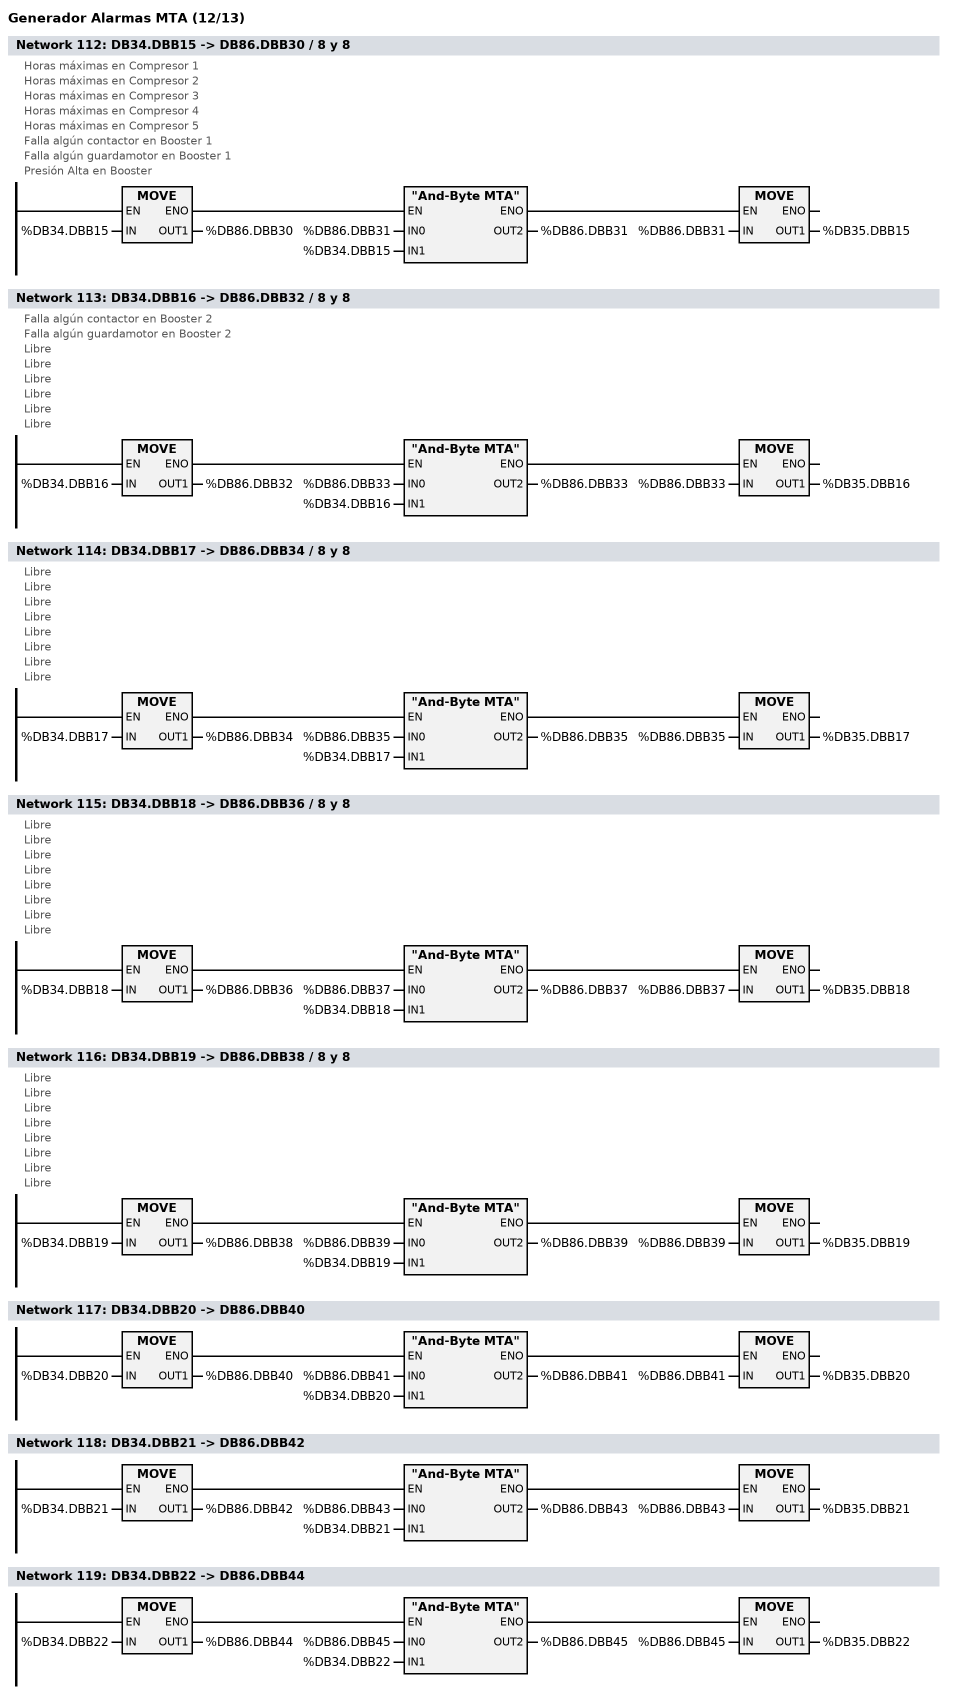
   RUNG wire#powerrail
      { S7_GenerateENO := "TRUE" } Move(in := %DB34.DBB15, out1 => %DB86.DBB30)
      "And-Byte MTA"(IN0 := %DB86.DBB31, IN1 := %DB34.DBB15, OUT2 => %DB86.DBB31)
      { S7_GenerateENO := "TRUE" } Move(in := %DB86.DBB31, out1 => %DB35.DBB15)
   END_RUNG
   // the same network as SCL:
   // ENO of a box is taken as its EN; it also drops when the box reports an error
   %DB86.DBB30 := %DB34.DBB15;
   "And-Byte MTA"(IN0 := %DB86.DBB31, IN1 := %DB34.DBB15, OUT2 => %DB86.DBB31, ENO => #_w1);
   IF #_w1 THEN %DB35.DBB15 := %DB86.DBB31; END_IF;
END_REGION

REGION Network 113: DB34.DBB16 -> DB86.DBB32 / 8 y 8
   // Falla algún contactor en Booster 2
   // Falla algún guardamotor en Booster 2
   // Libre
   // Libre
   // Libre
   // Libre
   // Libre
   // Libre
   RUNG wire#powerrail
      { S7_GenerateENO := "TRUE" } Move(in := %DB34.DBB16, out1 => %DB86.DBB32)
      "And-Byte MTA"(IN0 := %DB86.DBB33, IN1 := %DB34.DBB16, OUT2 => %DB86.DBB33)
      { S7_GenerateENO := "TRUE" } Move(in := %DB86.DBB33, out1 => %DB35.DBB16)
   END_RUNG
   // the same network as SCL:
   // ENO of a box is taken as its EN; it also drops when the box reports an error
   %DB86.DBB32 := %DB34.DBB16;
   "And-Byte MTA"(IN0 := %DB86.DBB33, IN1 := %DB34.DBB16, OUT2 => %DB86.DBB33, ENO => #_w1);
   IF #_w1 THEN %DB35.DBB16 := %DB86.DBB33; END_IF;
END_REGION

REGION Network 114: DB34.DBB17 -> DB86.DBB34 / 8 y 8
   // Libre
   // Libre
   // Libre
   // Libre
   // Libre
   // Libre
   // Libre
   // Libre
   RUNG wire#powerrail
      { S7_GenerateENO := "TRUE" } Move(in := %DB34.DBB17, out1 => %DB86.DBB34)
      "And-Byte MTA"(IN0 := %DB86.DBB35, IN1 := %DB34.DBB17, OUT2 => %DB86.DBB35)
      { S7_GenerateENO := "TRUE" } Move(in := %DB86.DBB35, out1 => %DB35.DBB17)
   END_RUNG
   // the same network as SCL:
   // ENO of a box is taken as its EN; it also drops when the box reports an error
   %DB86.DBB34 := %DB34.DBB17;
   "And-Byte MTA"(IN0 := %DB86.DBB35, IN1 := %DB34.DBB17, OUT2 => %DB86.DBB35, ENO => #_w1);
   IF #_w1 THEN %DB35.DBB17 := %DB86.DBB35; END_IF;
END_REGION

REGION Network 115: DB34.DBB18 -> DB86.DBB36 / 8 y 8
   // Libre
   // Libre
   // Libre
   // Libre
   // Libre
   // Libre
   // Libre
   // Libre
   RUNG wire#powerrail
      { S7_GenerateENO := "TRUE" } Move(in := %DB34.DBB18, out1 => %DB86.DBB36)
      "And-Byte MTA"(IN0 := %DB86.DBB37, IN1 := %DB34.DBB18, OUT2 => %DB86.DBB37)
      { S7_GenerateENO := "TRUE" } Move(in := %DB86.DBB37, out1 => %DB35.DBB18)
   END_RUNG
   // the same network as SCL:
   // ENO of a box is taken as its EN; it also drops when the box reports an error
   %DB86.DBB36 := %DB34.DBB18;
   "And-Byte MTA"(IN0 := %DB86.DBB37, IN1 := %DB34.DBB18, OUT2 => %DB86.DBB37, ENO => #_w1);
   IF #_w1 THEN %DB35.DBB18 := %DB86.DBB37; END_IF;
END_REGION

REGION Network 116: DB34.DBB19 -> DB86.DBB38 / 8 y 8
   // Libre
   // Libre
   // Libre
   // Libre
   // Libre
   // Libre
   // Libre
   // Libre
   RUNG wire#powerrail
      { S7_GenerateENO := "TRUE" } Move(in := %DB34.DBB19, out1 => %DB86.DBB38)
      "And-Byte MTA"(IN0 := %DB86.DBB39, IN1 := %DB34.DBB19, OUT2 => %DB86.DBB39)
      { S7_GenerateENO := "TRUE" } Move(in := %DB86.DBB39, out1 => %DB35.DBB19)
   END_RUNG
   // the same network as SCL:
   // ENO of a box is taken as its EN; it also drops when the box reports an error
   %DB86.DBB38 := %DB34.DBB19;
   "And-Byte MTA"(IN0 := %DB86.DBB39, IN1 := %DB34.DBB19, OUT2 => %DB86.DBB39, ENO => #_w1);
   IF #_w1 THEN %DB35.DBB19 := %DB86.DBB39; END_IF;
END_REGION

REGION Network 117: DB34.DBB20 -> DB86.DBB40
   RUNG wire#powerrail
      { S7_GenerateENO := "TRUE" } Move(in := %DB34.DBB20, out1 => %DB86.DBB40)
      "And-Byte MTA"(IN0 := %DB86.DBB41, IN1 := %DB34.DBB20, OUT2 => %DB86.DBB41)
      { S7_GenerateENO := "TRUE" } Move(in := %DB86.DBB41, out1 => %DB35.DBB20)
   END_RUNG
   // the same network as SCL:
   // ENO of a box is taken as its EN; it also drops when the box reports an error
   %DB86.DBB40 := %DB34.DBB20;
   "And-Byte MTA"(IN0 := %DB86.DBB41, IN1 := %DB34.DBB20, OUT2 => %DB86.DBB41, ENO => #_w1);
   IF #_w1 THEN %DB35.DBB20 := %DB86.DBB41; END_IF;
END_REGION

REGION Network 118: DB34.DBB21 -> DB86.DBB42
   RUNG wire#powerrail
      { S7_GenerateENO := "TRUE" } Move(in := %DB34.DBB21, out1 => %DB86.DBB42)
      "And-Byte MTA"(IN0 := %DB86.DBB43, IN1 := %DB34.DBB21, OUT2 => %DB86.DBB43)
      { S7_GenerateENO := "TRUE" } Move(in := %DB86.DBB43, out1 => %DB35.DBB21)
   END_RUNG
   // the same network as SCL:
   // ENO of a box is taken as its EN; it also drops when the box reports an error
   %DB86.DBB42 := %DB34.DBB21;
   "And-Byte MTA"(IN0 := %DB86.DBB43, IN1 := %DB34.DBB21, OUT2 => %DB86.DBB43, ENO => #_w1);
   IF #_w1 THEN %DB35.DBB21 := %DB86.DBB43; END_IF;
END_REGION

REGION Network 119: DB34.DBB22 -> DB86.DBB44
   RUNG wire#powerrail
      { S7_GenerateENO := "TRUE" } Move(in := %DB34.DBB22, out1 => %DB86.DBB44)
      "And-Byte MTA"(IN0 := %DB86.DBB45, IN1 := %DB34.DBB22, OUT2 => %DB86.DBB45)
      { S7_GenerateENO := "TRUE" } Move(in := %DB86.DBB45, out1 => %DB35.DBB22)
   END_RUNG
   // the same network as SCL:
   // ENO of a box is taken as its EN; it also drops when the box reports an error
   %DB86.DBB44 := %DB34.DBB22;
   "And-Byte MTA"(IN0 := %DB86.DBB45, IN1 := %DB34.DBB22, OUT2 => %DB86.DBB45, ENO => #_w1);
   IF #_w1 THEN %DB35.DBB22 := %DB86.DBB45; END_IF;
END_REGION

REGION Network 120: DB34.DBB23 -> DB86.DBB46
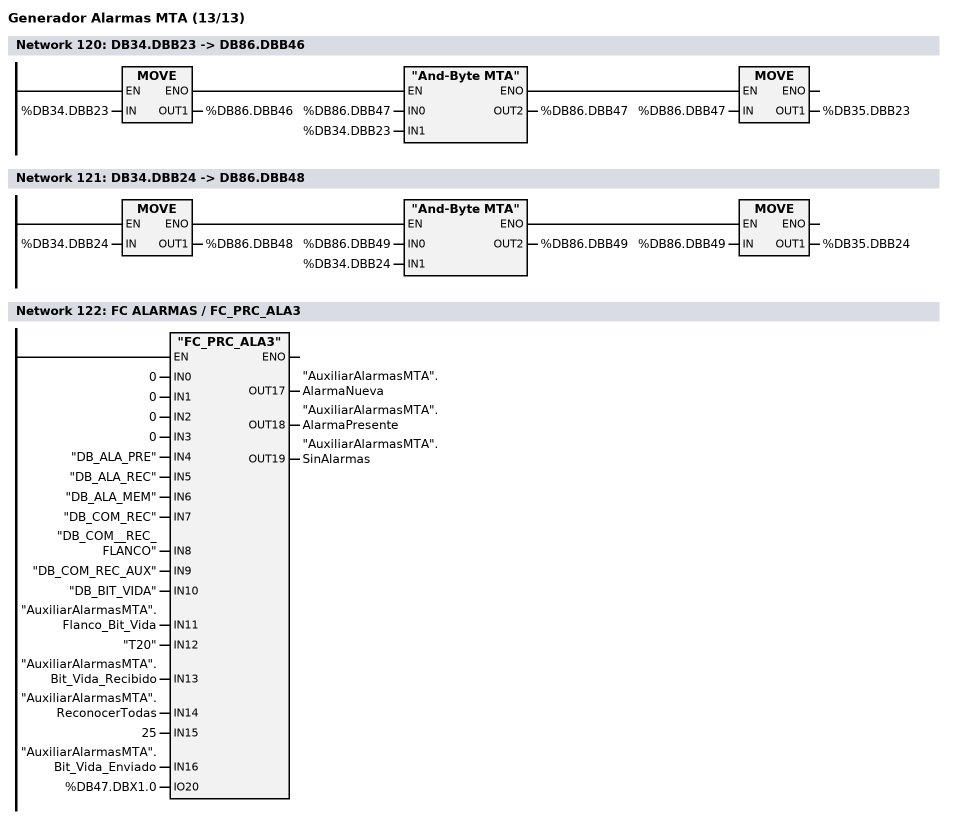
   RUNG wire#powerrail
      { S7_GenerateENO := "TRUE" } Move(in := %DB34.DBB23, out1 => %DB86.DBB46)
      "And-Byte MTA"(IN0 := %DB86.DBB47, IN1 := %DB34.DBB23, OUT2 => %DB86.DBB47)
      { S7_GenerateENO := "TRUE" } Move(in := %DB86.DBB47, out1 => %DB35.DBB23)
   END_RUNG
   // the same network as SCL:
   // ENO of a box is taken as its EN; it also drops when the box reports an error
   %DB86.DBB46 := %DB34.DBB23;
   "And-Byte MTA"(IN0 := %DB86.DBB47, IN1 := %DB34.DBB23, OUT2 => %DB86.DBB47, ENO => #_w1);
   IF #_w1 THEN %DB35.DBB23 := %DB86.DBB47; END_IF;
END_REGION

REGION Network 121: DB34.DBB24 -> DB86.DBB48
   RUNG wire#powerrail
      { S7_GenerateENO := "TRUE" } Move(in := %DB34.DBB24, out1 => %DB86.DBB48)
      "And-Byte MTA"(IN0 := %DB86.DBB49, IN1 := %DB34.DBB24, OUT2 => %DB86.DBB49)
      { S7_GenerateENO := "TRUE" } Move(in := %DB86.DBB49, out1 => %DB35.DBB24)
   END_RUNG
   // the same network as SCL:
   // ENO of a box is taken as its EN; it also drops when the box reports an error
   %DB86.DBB48 := %DB34.DBB24;
   "And-Byte MTA"(IN0 := %DB86.DBB49, IN1 := %DB34.DBB24, OUT2 => %DB86.DBB49, ENO => #_w1);
   IF #_w1 THEN %DB35.DBB24 := %DB86.DBB49; END_IF;
END_REGION

REGION Network 122: FC ALARMAS / FC_PRC_ALA3
   RUNG wire#powerrail
      "FC_PRC_ALA3"(IN0 := 0, IN1 := 0, IN2 := 0, IN3 := 0, IN4 := "DB_ALA_PRE", IN5 := "DB_ALA_REC", IN6 := "DB_ALA_MEM", IN7 := "DB_COM_REC", IN8 := "DB_COM__REC_FLANCO", IN9 := "DB_COM_REC_AUX", IN10 := "DB_BIT_VIDA", IN11 := "AuxiliarAlarmasMTA".Flanco_Bit_Vida, IN12 := "T20", IN13 := "AuxiliarAlarmasMTA".Bit_Vida_Recibido, IN14 := "AuxiliarAlarmasMTA".ReconocerTodas, IN15 := 25, IN16 := "AuxiliarAlarmasMTA".Bit_Vida_Enviado, IO20 := %DB47.DBX1.0, OUT17 => "AuxiliarAlarmasMTA".AlarmaNueva, OUT18 => "AuxiliarAlarmasMTA".AlarmaPresente, OUT19 => "AuxiliarAlarmasMTA".SinAlarmas)
   END_RUNG
   // the same network as SCL:
   "FC_PRC_ALA3"(IN0 := 0,
                 IN1 := 0,
                 IN2 := 0,
                 IN3 := 0,
                 IN4 := "DB_ALA_PRE",
                 IN5 := "DB_ALA_REC",
                 IN6 := "DB_ALA_MEM",
                 IN7 := "DB_COM_REC",
                 IN8 := "DB_COM__REC_FLANCO",
                 IN9 := "DB_COM_REC_AUX",
                 IN10 := "DB_BIT_VIDA",
                 IN11 := "AuxiliarAlarmasMTA".Flanco_Bit_Vida,
                 IN12 := "T20",
                 IN13 := "AuxiliarAlarmasMTA".Bit_Vida_Recibido,
                 IN14 := "AuxiliarAlarmasMTA".ReconocerTodas,
                 IN15 := 25,
                 IN16 := "AuxiliarAlarmasMTA".Bit_Vida_Enviado,
                 IO20 := %DB47.DBX1.0,
                 OUT17 => "AuxiliarAlarmasMTA".AlarmaNueva,
                 OUT18 => "AuxiliarAlarmasMTA".AlarmaPresente,
                 OUT19 => "AuxiliarAlarmasMTA".SinAlarmas);
END_REGION
END_FUNCTION

FUNCTION "FalCmpAlta" : Void   // FC49, LAD
{ S7_Optimized_Access := 'FALSE' }
VERSION : 0.1
BEGIN

REGION Network 1: Fallas de MC001 - Compresor de Alta ABC2
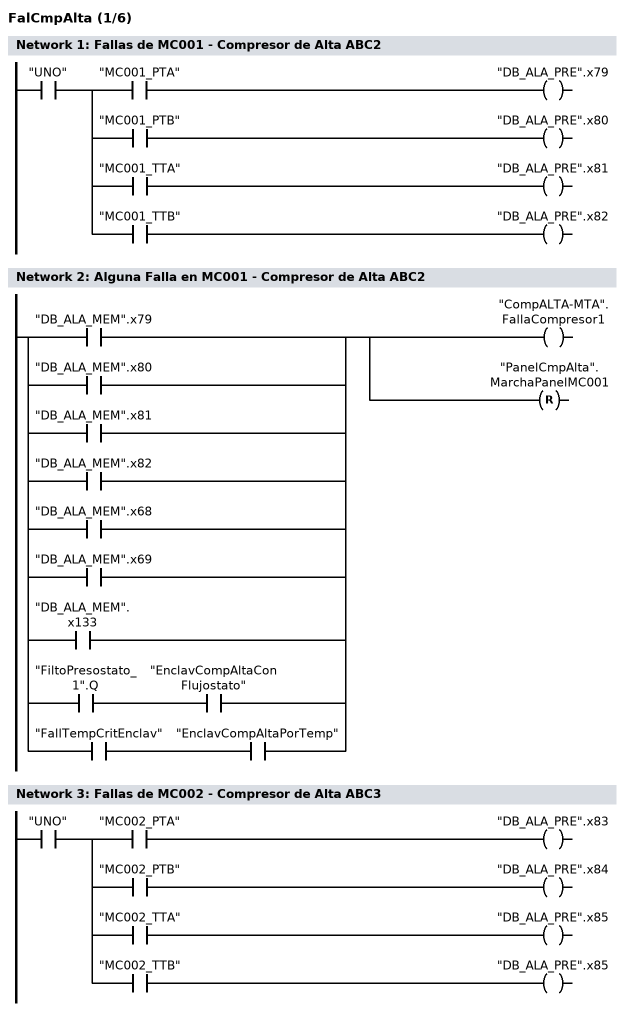
   RUNG wire#powerrail
      Contact( "UNO" )
      wire#w1
      Contact( "MC001_PTA" )
      Coil( "DB_ALA_PRE".x79 )
   END_RUNG
   RUNG wire#w1
      Contact( "MC001_PTB" )
      Coil( "DB_ALA_PRE".x80 )
   END_RUNG
   RUNG wire#w1
      Contact( "MC001_TTA" )
      Coil( "DB_ALA_PRE".x81 )
   END_RUNG
   RUNG wire#w1
      Contact( "MC001_TTB" )
      Coil( "DB_ALA_PRE".x82 )
   END_RUNG
   // the same network as SCL:
   "DB_ALA_PRE".x79 := "UNO" AND "MC001_PTA";
   "DB_ALA_PRE".x80 := "UNO" AND "MC001_PTB";
   "DB_ALA_PRE".x81 := "UNO" AND "MC001_TTA";
   "DB_ALA_PRE".x82 := "UNO" AND "MC001_TTB";
END_REGION

REGION Network 2: Alguna Falla en MC001 - Compresor de Alta ABC2
   RUNG wire#powerrail
      Contact( "DB_ALA_MEM".x79 )
      wire#w1
      Coil( "CompALTA-MTA".FallaCompresor1 )
   END_RUNG
   RUNG wire#powerrail
      Contact( "DB_ALA_MEM".x80 )
   END_RUNG wire#w1
   RUNG wire#powerrail
      Contact( "DB_ALA_MEM".x81 )
   END_RUNG wire#w1
   RUNG wire#powerrail
      Contact( "DB_ALA_MEM".x82 )
   END_RUNG wire#w1
   RUNG wire#powerrail
      Contact( "DB_ALA_MEM".x68 )
   END_RUNG wire#w1
   RUNG wire#powerrail
      Contact( "DB_ALA_MEM".x69 )
   END_RUNG wire#w1
   RUNG wire#powerrail
      Contact( "DB_ALA_MEM".x133 )
   END_RUNG wire#w1
   RUNG wire#powerrail
      Contact( "FiltoPresostato_1".Q )
      Contact( "EnclavCompAltaConFlujostato" )
   END_RUNG wire#w1
   RUNG wire#powerrail
      Contact( "FallTempCritEnclav" )
      Contact( "EnclavCompAltaPorTemp" )
   END_RUNG wire#w1
   RUNG wire#w1
      R_Coil( "PanelCmpAlta".MarchaPanelMC001 )
   END_RUNG
   // the same network as SCL:
   "CompALTA-MTA".FallaCompresor1 := "DB_ALA_MEM".x79 OR "DB_ALA_MEM".x80 OR "DB_ALA_MEM".x81 OR "DB_ALA_MEM".x82 OR "DB_ALA_MEM".x68 OR "DB_ALA_MEM".x69 OR "DB_ALA_MEM".x133 OR ("FiltoPresostato_1".Q AND "EnclavCompAltaConFlujostato") OR ("FallTempCritEnclav" AND "EnclavCompAltaPorTemp");
   IF "CompALTA-MTA".FallaCompresor1 THEN "PanelCmpAlta".MarchaPanelMC001 := FALSE; END_IF;
END_REGION

REGION Network 3: Fallas de MC002 - Compresor de Alta ABC3
   RUNG wire#powerrail
      Contact( "UNO" )
      wire#w1
      Contact( "MC002_PTA" )
      Coil( "DB_ALA_PRE".x83 )
   END_RUNG
   RUNG wire#w1
      Contact( "MC002_PTB" )
      Coil( "DB_ALA_PRE".x84 )
   END_RUNG
   RUNG wire#w1
      Contact( "MC002_TTA" )
      Coil( "DB_ALA_PRE".x85 )
   END_RUNG
   RUNG wire#w1
      Contact( "MC002_TTB" )
      Coil( "DB_ALA_PRE".x85 )
   END_RUNG
   // the same network as SCL:
   "DB_ALA_PRE".x83 := "UNO" AND "MC002_PTA";
   "DB_ALA_PRE".x84 := "UNO" AND "MC002_PTB";
   "DB_ALA_PRE".x85 := "UNO" AND "MC002_TTA";
   "DB_ALA_PRE".x85 := "UNO" AND "MC002_TTB";
END_REGION

REGION Network 4: Alguna Falla en MC002 - Compresor de Alta ABC3
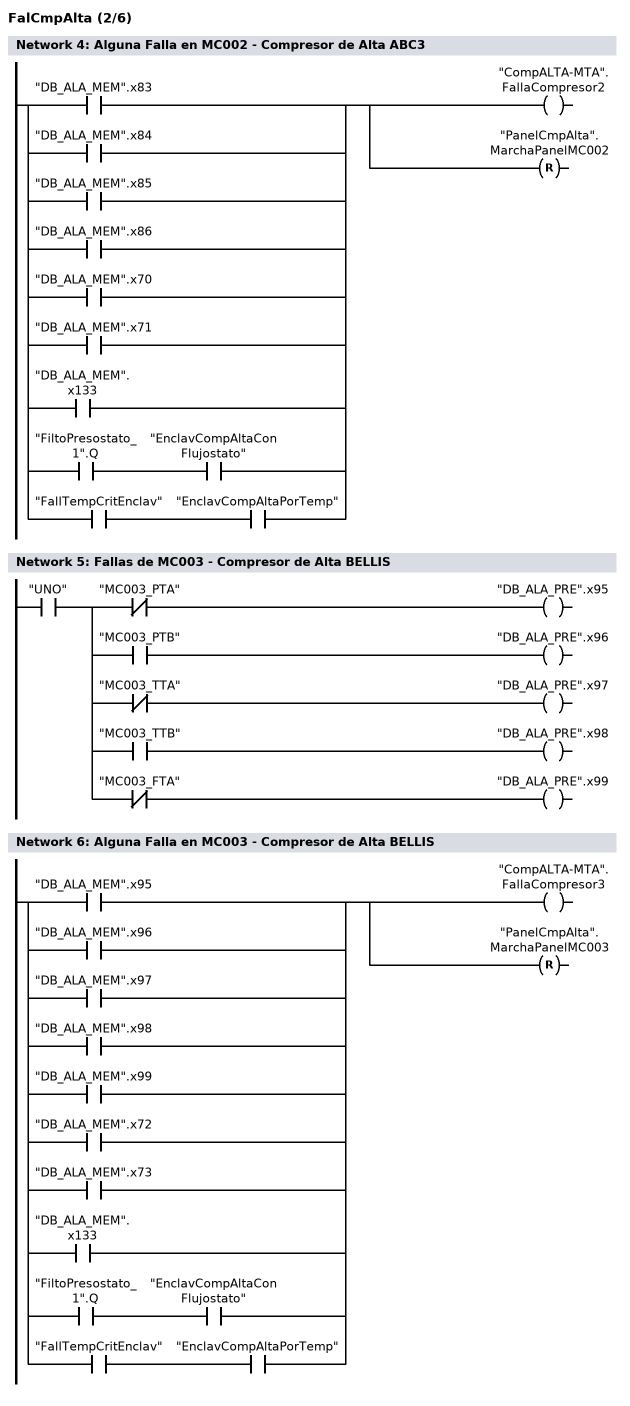
   RUNG wire#powerrail
      Contact( "DB_ALA_MEM".x83 )
      wire#w1
      Coil( "CompALTA-MTA".FallaCompresor2 )
   END_RUNG
   RUNG wire#powerrail
      Contact( "DB_ALA_MEM".x84 )
   END_RUNG wire#w1
   RUNG wire#powerrail
      Contact( "DB_ALA_MEM".x85 )
   END_RUNG wire#w1
   RUNG wire#powerrail
      Contact( "DB_ALA_MEM".x86 )
   END_RUNG wire#w1
   RUNG wire#powerrail
      Contact( "DB_ALA_MEM".x70 )
   END_RUNG wire#w1
   RUNG wire#powerrail
      Contact( "DB_ALA_MEM".x71 )
   END_RUNG wire#w1
   RUNG wire#powerrail
      Contact( "DB_ALA_MEM".x133 )
   END_RUNG wire#w1
   RUNG wire#powerrail
      Contact( "FiltoPresostato_1".Q )
      Contact( "EnclavCompAltaConFlujostato" )
   END_RUNG wire#w1
   RUNG wire#powerrail
      Contact( "FallTempCritEnclav" )
      Contact( "EnclavCompAltaPorTemp" )
   END_RUNG wire#w1
   RUNG wire#w1
      R_Coil( "PanelCmpAlta".MarchaPanelMC002 )
   END_RUNG
   // the same network as SCL:
   "CompALTA-MTA".FallaCompresor2 := "DB_ALA_MEM".x83 OR "DB_ALA_MEM".x84 OR "DB_ALA_MEM".x85 OR "DB_ALA_MEM".x86 OR "DB_ALA_MEM".x70 OR "DB_ALA_MEM".x71 OR "DB_ALA_MEM".x133 OR ("FiltoPresostato_1".Q AND "EnclavCompAltaConFlujostato") OR ("FallTempCritEnclav" AND "EnclavCompAltaPorTemp");
   IF "CompALTA-MTA".FallaCompresor2 THEN "PanelCmpAlta".MarchaPanelMC002 := FALSE; END_IF;
END_REGION

REGION Network 5: Fallas de MC003 - Compresor de Alta BELLIS
   RUNG wire#powerrail
      Contact( "UNO" )
      wire#w1
      I_Contact( "MC003_PTA" )
      Coil( "DB_ALA_PRE".x95 )
   END_RUNG
   RUNG wire#w1
      Contact( "MC003_PTB" )
      Coil( "DB_ALA_PRE".x96 )
   END_RUNG
   RUNG wire#w1
      I_Contact( "MC003_TTA" )
      Coil( "DB_ALA_PRE".x97 )
   END_RUNG
   RUNG wire#w1
      Contact( "MC003_TTB" )
      Coil( "DB_ALA_PRE".x98 )
   END_RUNG
   RUNG wire#w1
      I_Contact( "MC003_FTA" )
      Coil( "DB_ALA_PRE".x99 )
   END_RUNG
   // the same network as SCL:
   "DB_ALA_PRE".x95 := "UNO" AND NOT "MC003_PTA";
   "DB_ALA_PRE".x96 := "UNO" AND "MC003_PTB";
   "DB_ALA_PRE".x97 := "UNO" AND NOT "MC003_TTA";
   "DB_ALA_PRE".x98 := "UNO" AND "MC003_TTB";
   "DB_ALA_PRE".x99 := "UNO" AND NOT "MC003_FTA";
END_REGION

REGION Network 6: Alguna Falla en MC003 - Compresor de Alta BELLIS
   RUNG wire#powerrail
      Contact( "DB_ALA_MEM".x95 )
      wire#w1
      Coil( "CompALTA-MTA".FallaCompresor3 )
   END_RUNG
   RUNG wire#powerrail
      Contact( "DB_ALA_MEM".x96 )
   END_RUNG wire#w1
   RUNG wire#powerrail
      Contact( "DB_ALA_MEM".x97 )
   END_RUNG wire#w1
   RUNG wire#powerrail
      Contact( "DB_ALA_MEM".x98 )
   END_RUNG wire#w1
   RUNG wire#powerrail
      Contact( "DB_ALA_MEM".x99 )
   END_RUNG wire#w1
   RUNG wire#powerrail
      Contact( "DB_ALA_MEM".x72 )
   END_RUNG wire#w1
   RUNG wire#powerrail
      Contact( "DB_ALA_MEM".x73 )
   END_RUNG wire#w1
   RUNG wire#powerrail
      Contact( "DB_ALA_MEM".x133 )
   END_RUNG wire#w1
   RUNG wire#powerrail
      Contact( "FiltoPresostato_1".Q )
      Contact( "EnclavCompAltaConFlujostato" )
   END_RUNG wire#w1
   RUNG wire#powerrail
      Contact( "FallTempCritEnclav" )
      Contact( "EnclavCompAltaPorTemp" )
   END_RUNG wire#w1
   RUNG wire#w1
      R_Coil( "PanelCmpAlta".MarchaPanelMC003 )
   END_RUNG
   // the same network as SCL:
   "CompALTA-MTA".FallaCompresor3 := "DB_ALA_MEM".x95 OR "DB_ALA_MEM".x96 OR "DB_ALA_MEM".x97 OR "DB_ALA_MEM".x98 OR "DB_ALA_MEM".x99 OR "DB_ALA_MEM".x72 OR "DB_ALA_MEM".x73 OR "DB_ALA_MEM".x133 OR ("FiltoPresostato_1".Q AND "EnclavCompAltaConFlujostato") OR ("FallTempCritEnclav" AND "EnclavCompAltaPorTemp");
   IF "CompALTA-MTA".FallaCompresor3 THEN "PanelCmpAlta".MarchaPanelMC003 := FALSE; END_IF;
END_REGION

REGION Network 7: Fallas de MC004 - Compresor de Alta ABC4
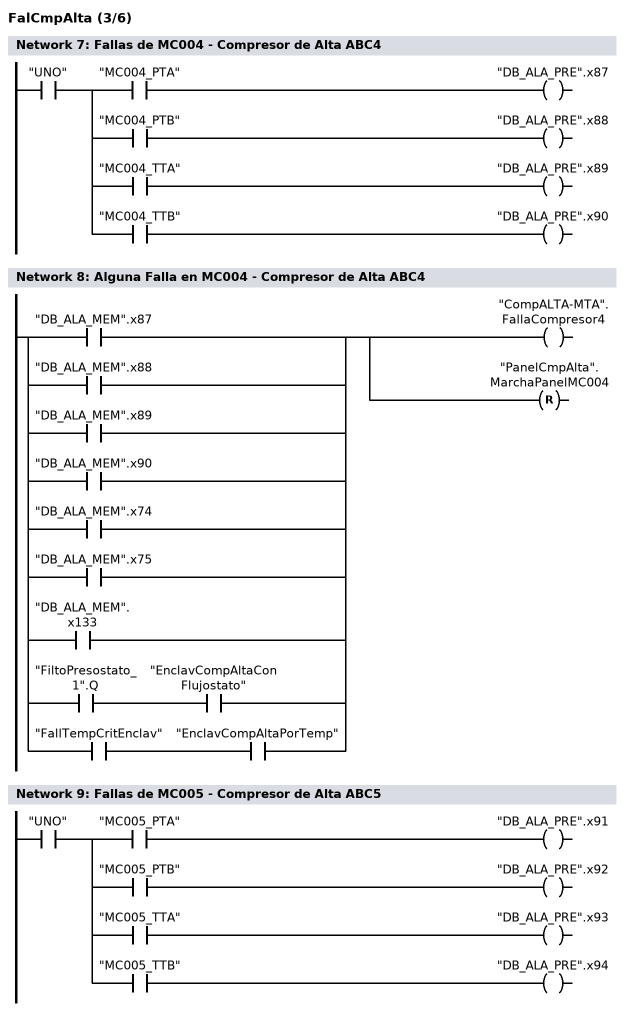
   RUNG wire#powerrail
      Contact( "UNO" )
      wire#w1
      Contact( "MC004_PTA" )
      Coil( "DB_ALA_PRE".x87 )
   END_RUNG
   RUNG wire#w1
      Contact( "MC004_PTB" )
      Coil( "DB_ALA_PRE".x88 )
   END_RUNG
   RUNG wire#w1
      Contact( "MC004_TTA" )
      Coil( "DB_ALA_PRE".x89 )
   END_RUNG
   RUNG wire#w1
      Contact( "MC004_TTB" )
      Coil( "DB_ALA_PRE".x90 )
   END_RUNG
   // the same network as SCL:
   "DB_ALA_PRE".x87 := "UNO" AND "MC004_PTA";
   "DB_ALA_PRE".x88 := "UNO" AND "MC004_PTB";
   "DB_ALA_PRE".x89 := "UNO" AND "MC004_TTA";
   "DB_ALA_PRE".x90 := "UNO" AND "MC004_TTB";
END_REGION

REGION Network 8: Alguna Falla en MC004 - Compresor de Alta ABC4
   RUNG wire#powerrail
      Contact( "DB_ALA_MEM".x87 )
      wire#w1
      Coil( "CompALTA-MTA".FallaCompresor4 )
   END_RUNG
   RUNG wire#powerrail
      Contact( "DB_ALA_MEM".x88 )
   END_RUNG wire#w1
   RUNG wire#powerrail
      Contact( "DB_ALA_MEM".x89 )
   END_RUNG wire#w1
   RUNG wire#powerrail
      Contact( "DB_ALA_MEM".x90 )
   END_RUNG wire#w1
   RUNG wire#powerrail
      Contact( "DB_ALA_MEM".x74 )
   END_RUNG wire#w1
   RUNG wire#powerrail
      Contact( "DB_ALA_MEM".x75 )
   END_RUNG wire#w1
   RUNG wire#powerrail
      Contact( "DB_ALA_MEM".x133 )
   END_RUNG wire#w1
   RUNG wire#powerrail
      Contact( "FiltoPresostato_1".Q )
      Contact( "EnclavCompAltaConFlujostato" )
   END_RUNG wire#w1
   RUNG wire#powerrail
      Contact( "FallTempCritEnclav" )
      Contact( "EnclavCompAltaPorTemp" )
   END_RUNG wire#w1
   RUNG wire#w1
      R_Coil( "PanelCmpAlta".MarchaPanelMC004 )
   END_RUNG
   // the same network as SCL:
   "CompALTA-MTA".FallaCompresor4 := "DB_ALA_MEM".x87 OR "DB_ALA_MEM".x88 OR "DB_ALA_MEM".x89 OR "DB_ALA_MEM".x90 OR "DB_ALA_MEM".x74 OR "DB_ALA_MEM".x75 OR "DB_ALA_MEM".x133 OR ("FiltoPresostato_1".Q AND "EnclavCompAltaConFlujostato") OR ("FallTempCritEnclav" AND "EnclavCompAltaPorTemp");
   IF "CompALTA-MTA".FallaCompresor4 THEN "PanelCmpAlta".MarchaPanelMC004 := FALSE; END_IF;
END_REGION

REGION Network 9: Fallas de MC005 - Compresor de Alta ABC5
   RUNG wire#powerrail
      Contact( "UNO" )
      wire#w1
      Contact( "MC005_PTA" )
      Coil( "DB_ALA_PRE".x91 )
   END_RUNG
   RUNG wire#w1
      Contact( "MC005_PTB" )
      Coil( "DB_ALA_PRE".x92 )
   END_RUNG
   RUNG wire#w1
      Contact( "MC005_TTA" )
      Coil( "DB_ALA_PRE".x93 )
   END_RUNG
   RUNG wire#w1
      Contact( "MC005_TTB" )
      Coil( "DB_ALA_PRE".x94 )
   END_RUNG
   // the same network as SCL:
   "DB_ALA_PRE".x91 := "UNO" AND "MC005_PTA";
   "DB_ALA_PRE".x92 := "UNO" AND "MC005_PTB";
   "DB_ALA_PRE".x93 := "UNO" AND "MC005_TTA";
   "DB_ALA_PRE".x94 := "UNO" AND "MC005_TTB";
END_REGION

REGION Network 10: Alguna Falla en MC005 - Compresor de Alta ABC5
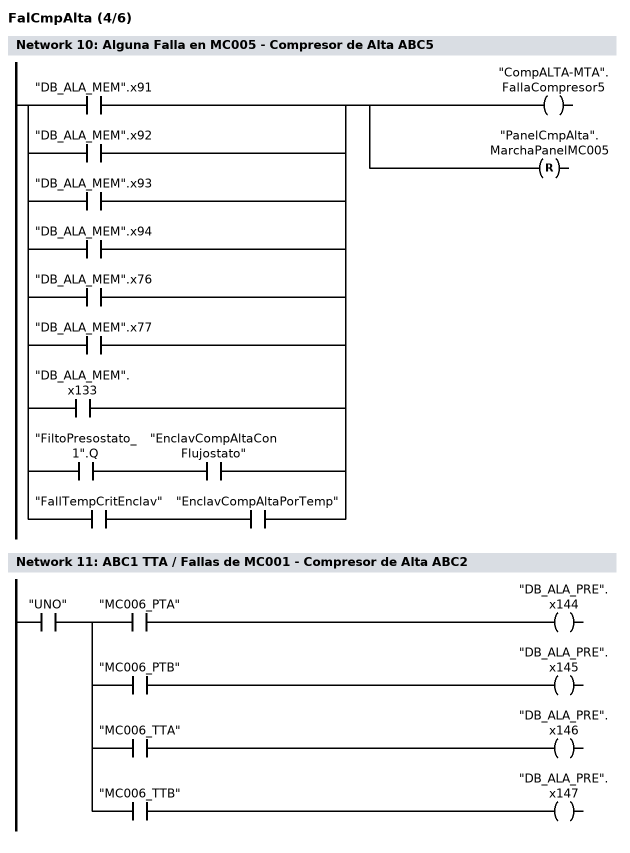
   RUNG wire#powerrail
      Contact( "DB_ALA_MEM".x91 )
      wire#w1
      Coil( "CompALTA-MTA".FallaCompresor5 )
   END_RUNG
   RUNG wire#powerrail
      Contact( "DB_ALA_MEM".x92 )
   END_RUNG wire#w1
   RUNG wire#powerrail
      Contact( "DB_ALA_MEM".x93 )
   END_RUNG wire#w1
   RUNG wire#powerrail
      Contact( "DB_ALA_MEM".x94 )
   END_RUNG wire#w1
   RUNG wire#powerrail
      Contact( "DB_ALA_MEM".x76 )
   END_RUNG wire#w1
   RUNG wire#powerrail
      Contact( "DB_ALA_MEM".x77 )
   END_RUNG wire#w1
   RUNG wire#powerrail
      Contact( "DB_ALA_MEM".x133 )
   END_RUNG wire#w1
   RUNG wire#powerrail
      Contact( "FiltoPresostato_1".Q )
      Contact( "EnclavCompAltaConFlujostato" )
   END_RUNG wire#w1
   RUNG wire#powerrail
      Contact( "FallTempCritEnclav" )
      Contact( "EnclavCompAltaPorTemp" )
   END_RUNG wire#w1
   RUNG wire#w1
      R_Coil( "PanelCmpAlta".MarchaPanelMC005 )
   END_RUNG
   // the same network as SCL:
   "CompALTA-MTA".FallaCompresor5 := "DB_ALA_MEM".x91 OR "DB_ALA_MEM".x92 OR "DB_ALA_MEM".x93 OR "DB_ALA_MEM".x94 OR "DB_ALA_MEM".x76 OR "DB_ALA_MEM".x77 OR "DB_ALA_MEM".x133 OR ("FiltoPresostato_1".Q AND "EnclavCompAltaConFlujostato") OR ("FallTempCritEnclav" AND "EnclavCompAltaPorTemp");
   IF "CompALTA-MTA".FallaCompresor5 THEN "PanelCmpAlta".MarchaPanelMC005 := FALSE; END_IF;
END_REGION

REGION Network 11: ABC1 TTA / Fallas de MC001 - Compresor de Alta ABC2
   RUNG wire#powerrail
      Contact( "UNO" )
      wire#w1
      Contact( "MC006_PTA" )
      Coil( "DB_ALA_PRE".x144 )
   END_RUNG
   RUNG wire#w1
      Contact( "MC006_PTB" )
      Coil( "DB_ALA_PRE".x145 )
   END_RUNG
   RUNG wire#w1
      Contact( "MC006_TTA" )
      Coil( "DB_ALA_PRE".x146 )
   END_RUNG
   RUNG wire#w1
      Contact( "MC006_TTB" )
      Coil( "DB_ALA_PRE".x147 )
   END_RUNG
   // the same network as SCL:
   "DB_ALA_PRE".x144 := "UNO" AND "MC006_PTA";
   "DB_ALA_PRE".x145 := "UNO" AND "MC006_PTB";
   "DB_ALA_PRE".x146 := "UNO" AND "MC006_TTA";
   "DB_ALA_PRE".x147 := "UNO" AND "MC006_TTB";
END_REGION

REGION Network 12: Alguna Falla en MC001 - Compresor de Alta ABC2
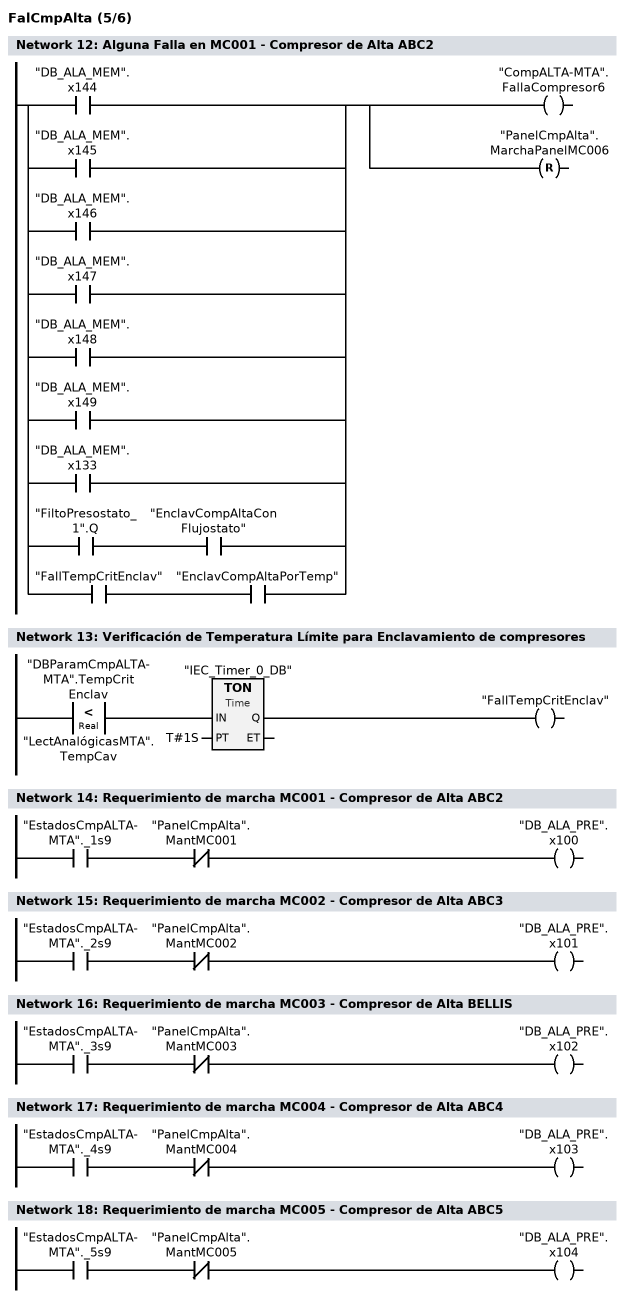
   RUNG wire#powerrail
      Contact( "DB_ALA_MEM".x144 )
      wire#w1
      Coil( "CompALTA-MTA".FallaCompresor6 )
   END_RUNG
   RUNG wire#powerrail
      Contact( "DB_ALA_MEM".x145 )
   END_RUNG wire#w1
   RUNG wire#powerrail
      Contact( "DB_ALA_MEM".x146 )
   END_RUNG wire#w1
   RUNG wire#powerrail
      Contact( "DB_ALA_MEM".x147 )
   END_RUNG wire#w1
   RUNG wire#powerrail
      Contact( "DB_ALA_MEM".x148 )
   END_RUNG wire#w1
   RUNG wire#powerrail
      Contact( "DB_ALA_MEM".x149 )
   END_RUNG wire#w1
   RUNG wire#powerrail
      Contact( "DB_ALA_MEM".x133 )
   END_RUNG wire#w1
   RUNG wire#powerrail
      Contact( "FiltoPresostato_1".Q )
      Contact( "EnclavCompAltaConFlujostato" )
   END_RUNG wire#w1
   RUNG wire#powerrail
      Contact( "FallTempCritEnclav" )
      Contact( "EnclavCompAltaPorTemp" )
   END_RUNG wire#w1
   RUNG wire#w1
      R_Coil( "PanelCmpAlta".MarchaPanelMC006 )
   END_RUNG
   // the same network as SCL:
   "CompALTA-MTA".FallaCompresor6 := "DB_ALA_MEM".x144 OR "DB_ALA_MEM".x145 OR "DB_ALA_MEM".x146 OR "DB_ALA_MEM".x147 OR "DB_ALA_MEM".x148 OR "DB_ALA_MEM".x149 OR "DB_ALA_MEM".x133 OR ("FiltoPresostato_1".Q AND "EnclavCompAltaConFlujostato") OR ("FallTempCritEnclav" AND "EnclavCompAltaPorTemp");
   IF "CompALTA-MTA".FallaCompresor6 THEN "PanelCmpAlta".MarchaPanelMC006 := FALSE; END_IF;
END_REGION

REGION Network 13: Verificación de Temperatura Límite para Enclavamiento de compresores
   "IEC_Timer_0_DB".TON(IN := "DBParamCmpALTA-MTA".TempCritEnclav < "LectAnalógicasMTA".TempCav, PT := T#1S);
   "FallTempCritEnclav" := "IEC_Timer_0_DB".Q;
END_REGION

REGION Network 14: Requerimiento de marcha MC001 - Compresor de Alta ABC2
   RUNG wire#powerrail
      Contact( "EstadosCmpALTA-MTA"._1s9 )
      I_Contact( "PanelCmpAlta".MantMC001 )
      Coil( "DB_ALA_PRE".x100 )
   END_RUNG
   // the same network as SCL:
   "DB_ALA_PRE".x100 := "EstadosCmpALTA-MTA"._1s9 AND NOT "PanelCmpAlta".MantMC001;
END_REGION

REGION Network 15: Requerimiento de marcha MC002 - Compresor de Alta ABC3
   RUNG wire#powerrail
      Contact( "EstadosCmpALTA-MTA"._2s9 )
      I_Contact( "PanelCmpAlta".MantMC002 )
      Coil( "DB_ALA_PRE".x101 )
   END_RUNG
   // the same network as SCL:
   "DB_ALA_PRE".x101 := "EstadosCmpALTA-MTA"._2s9 AND NOT "PanelCmpAlta".MantMC002;
END_REGION

REGION Network 16: Requerimiento de marcha MC003 - Compresor de Alta BELLIS
   RUNG wire#powerrail
      Contact( "EstadosCmpALTA-MTA"._3s9 )
      I_Contact( "PanelCmpAlta".MantMC003 )
      Coil( "DB_ALA_PRE".x102 )
   END_RUNG
   // the same network as SCL:
   "DB_ALA_PRE".x102 := "EstadosCmpALTA-MTA"._3s9 AND NOT "PanelCmpAlta".MantMC003;
END_REGION

REGION Network 17: Requerimiento de marcha MC004 - Compresor de Alta ABC4
   RUNG wire#powerrail
      Contact( "EstadosCmpALTA-MTA"._4s9 )
      I_Contact( "PanelCmpAlta".MantMC004 )
      Coil( "DB_ALA_PRE".x103 )
   END_RUNG
   // the same network as SCL:
   "DB_ALA_PRE".x103 := "EstadosCmpALTA-MTA"._4s9 AND NOT "PanelCmpAlta".MantMC004;
END_REGION

REGION Network 18: Requerimiento de marcha MC005 - Compresor de Alta ABC5
   RUNG wire#powerrail
      Contact( "EstadosCmpALTA-MTA"._5s9 )
      I_Contact( "PanelCmpAlta".MantMC005 )
      Coil( "DB_ALA_PRE".x104 )
   END_RUNG
   // the same network as SCL:
   "DB_ALA_PRE".x104 := "EstadosCmpALTA-MTA"._5s9 AND NOT "PanelCmpAlta".MantMC005;
END_REGION

REGION Network 19: Requerimiento de marcha MC001 - Compresor de Alta ABC2
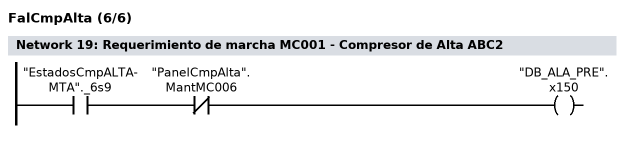
   RUNG wire#powerrail
      Contact( "EstadosCmpALTA-MTA"._6s9 )
      I_Contact( "PanelCmpAlta".MantMC006 )
      Coil( "DB_ALA_PRE".x150 )
   END_RUNG
   // the same network as SCL:
   "DB_ALA_PRE".x150 := "EstadosCmpALTA-MTA"._6s9 AND NOT "PanelCmpAlta".MantMC006;
END_REGION
END_FUNCTION

// folder: Auxiliares

FUNCTION "AjusteEntrada-SalidaMTA" : Void   // FC6, LAD
{ S7_Optimized_Access := 'FALSE' }
VERSION : 0.1
BEGIN

REGION Network 1
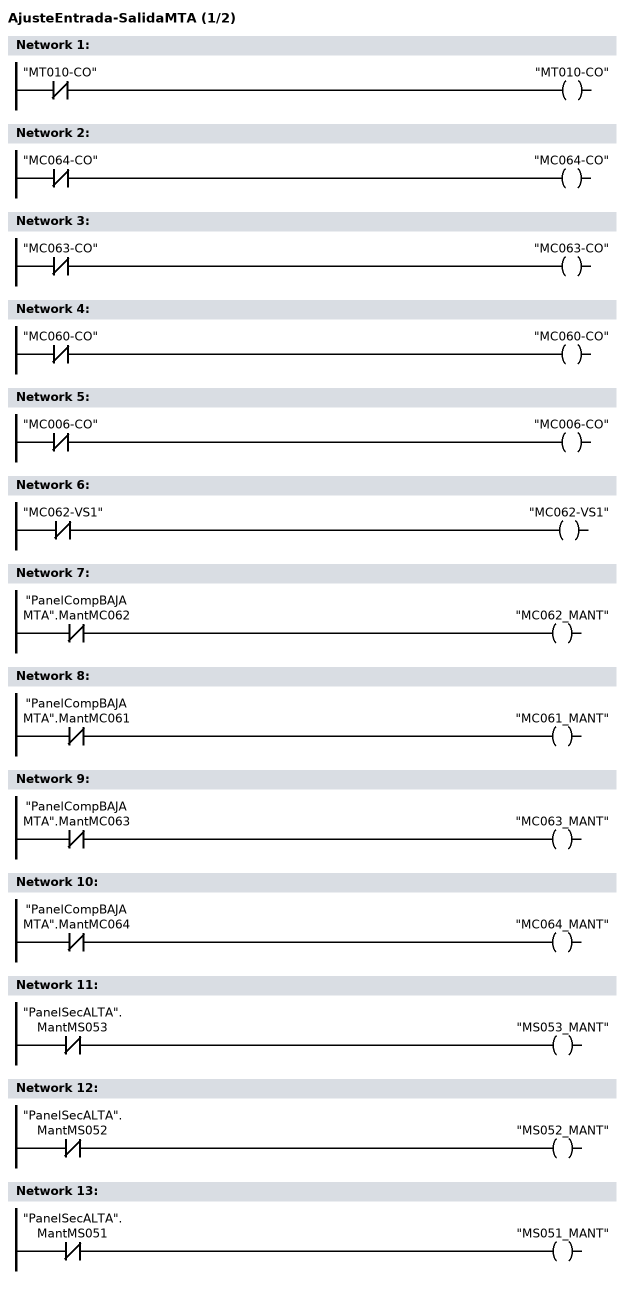
   RUNG wire#powerrail
      I_Contact( "MT010-CO" )
      Coil( "MT010-CO" )
   END_RUNG
   // the same network as SCL:
   "MT010-CO" := NOT "MT010-CO";
END_REGION

REGION Network 2
   RUNG wire#powerrail
      I_Contact( "MC064-CO" )
      Coil( "MC064-CO" )
   END_RUNG
   // the same network as SCL:
   "MC064-CO" := NOT "MC064-CO";
END_REGION

REGION Network 3
   RUNG wire#powerrail
      I_Contact( "MC063-CO" )
      Coil( "MC063-CO" )
   END_RUNG
   // the same network as SCL:
   "MC063-CO" := NOT "MC063-CO";
END_REGION

REGION Network 4
   RUNG wire#powerrail
      I_Contact( "MC060-CO" )
      Coil( "MC060-CO" )
   END_RUNG
   // the same network as SCL:
   "MC060-CO" := NOT "MC060-CO";
END_REGION

REGION Network 5
   RUNG wire#powerrail
      I_Contact( "MC006-CO" )
      Coil( "MC006-CO" )
   END_RUNG
   // the same network as SCL:
   "MC006-CO" := NOT "MC006-CO";
END_REGION

REGION Network 6
   RUNG wire#powerrail
      I_Contact( "MC062-VS1" )
      Coil( "MC062-VS1" )
   END_RUNG
   // the same network as SCL:
   "MC062-VS1" := NOT "MC062-VS1";
END_REGION

REGION Network 7
   RUNG wire#powerrail
      I_Contact( "PanelCompBAJA MTA".MantMC062 )
      Coil( "MC062_MANT" )
   END_RUNG
   // the same network as SCL:
   "MC062_MANT" := NOT "PanelCompBAJA MTA".MantMC062;
END_REGION

REGION Network 8
   RUNG wire#powerrail
      I_Contact( "PanelCompBAJA MTA".MantMC061 )
      Coil( "MC061_MANT" )
   END_RUNG
   // the same network as SCL:
   "MC061_MANT" := NOT "PanelCompBAJA MTA".MantMC061;
END_REGION

REGION Network 9
   RUNG wire#powerrail
      I_Contact( "PanelCompBAJA MTA".MantMC063 )
      Coil( "MC063_MANT" )
   END_RUNG
   // the same network as SCL:
   "MC063_MANT" := NOT "PanelCompBAJA MTA".MantMC063;
END_REGION

REGION Network 10
   RUNG wire#powerrail
      I_Contact( "PanelCompBAJA MTA".MantMC064 )
      Coil( "MC064_MANT" )
   END_RUNG
   // the same network as SCL:
   "MC064_MANT" := NOT "PanelCompBAJA MTA".MantMC064;
END_REGION

REGION Network 11
   RUNG wire#powerrail
      I_Contact( "PanelSecALTA".MantMS053 )
      Coil( "MS053_MANT" )
   END_RUNG
   // the same network as SCL:
   "MS053_MANT" := NOT "PanelSecALTA".MantMS053;
END_REGION

REGION Network 12
   RUNG wire#powerrail
      I_Contact( "PanelSecALTA".MantMS052 )
      Coil( "MS052_MANT" )
   END_RUNG
   // the same network as SCL:
   "MS052_MANT" := NOT "PanelSecALTA".MantMS052;
END_REGION

REGION Network 13
   RUNG wire#powerrail
      I_Contact( "PanelSecALTA".MantMS051 )
      Coil( "MS051_MANT" )
   END_RUNG
   // the same network as SCL:
   "MS051_MANT" := NOT "PanelSecALTA".MantMS051;
END_REGION

REGION Network 14
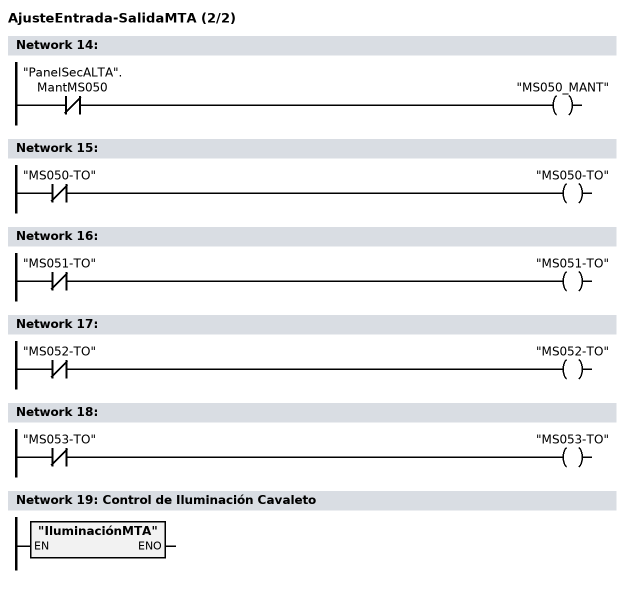
   RUNG wire#powerrail
      I_Contact( "PanelSecALTA".MantMS050 )
      Coil( "MS050_MANT" )
   END_RUNG
   // the same network as SCL:
   "MS050_MANT" := NOT "PanelSecALTA".MantMS050;
END_REGION
